
           REGION "SEND TO HMI"
               #saveAct := #partCall.row[#i].pbSelection.actuate;
               #partCall.row[#i] := #requests.row[#pRow];
               #partCall.row[#i].pbSelection.actuate := #saveAct;
           END_REGION

       END_FOR;
   END_REGION
END_FUNCTION_BLOCK

FUNCTION_BLOCK "Clear Part Requests"   // FB17, SCL
{ S7_Optimized_Access := 'TRUE' }
VERSION : 0.1
   VAR_INPUT
      clearRequest : Bool;
   END_VAR
   VAR_IN_OUT
      requests : "Part Request Data";
      partCall : "Part Call Screen";
      currentRowCount : Int;
   END_VAR
   VAR_TEMP
      blankRow : "Table Row";
      i : Int;
      maxRows : Int;
   END_VAR
BEGIN
   REGION "ON REQUEST"
       IF #clearRequest THEN

           REGION "HMI TABLE"

               REGION "COPY TO LOCAL"
                   #maxRows := "partReqHmiRowCount";
               END_REGION

               REGION "CLEAR ROWS"
                   FOR #i := 0 TO #maxRows DO
                       #partCall.row[#i] := #blankRow;
                   END_FOR;
               END_REGION

           END_REGION

           REGION "PART REQUEST DATA BASE"

               REGION "COPY TO LOCAL"
                   #maxRows := "partReqDataRowCount";
               END_REGION

               REGION "CLEAR ROWS"
                   FOR #i := 0 TO #maxRows DO
                       #requests.row[#i] := #blankRow;
                       #currentRowCount := 0;
                   END_FOR;
               END_REGION

           END_REGION

       END_IF;
   END_REGION
END_FUNCTION_BLOCK

FUNCTION_BLOCK "Load Default Timer Presets"   // FB18, SCL
{ S7_Optimized_Access := 'TRUE' }
VERSION : 0.1
   VAR_INPUT
      req : Bool;
   END_VAR
   VAR_IN_OUT
      stations : "Stations";
   END_VAR
   VAR
      oldReq : Bool;
   END_VAR
   VAR_TEMP
      alotted : Real;
      btnCount : Int;
      critical : Real;
      i : Int;
      j : Int;
      partNumber : WString;
      stnCount : Int;
      tmrReal : Real;
   END_VAR
BEGIN
   REGION "COPY TO LOCAL"
       #alotted := "defaultAlotted";
       #btnCount := "ptsPerStn";
       #critical := "defaultCritical";
       #stnCount := #stnCount;
   END_REGION

   REGION "ON REQUEST RISING EDGE"
       IF #req AND NOT #oldReq THEN

           REGION "LOOP THROUGH STATIONS" 
               FOR #i := 0 TO #stnCount DO

                   REGION "LOOP THROUGH BUTTONS"
                       FOR #j := 0 TO #btnCount DO

                           REGION "COPY TO LOCAL"
                               #partNumber := #stations.me[#i].partNumbers[#j];
                           END_REGION

                           REGION "IF BUTTON HAS ASSOCIATED PN"
                               IF LEN(#partNumber) <> 0 THEN

                                   REGION "COPY TO LOCAL"
                                       #tmrReal := #stations.me[#i].presetTime.allotted[#j];
                                   END_REGION

                                   REGION "ON NO TIME ENTERED"
                                       IF #tmrReal = 0.0 THEN

                                           REGION "ASSIGN ALLOTTED VALUES"
                                               #stations.me[#i].presetTime.allotted[#j] := #alotted;
                                           END_REGION

                                       END_IF;
                                   END_REGION

                                   REGION "COPY TO LOCAL"
                                       #tmrReal := #stations.me[#i].presetTime.critical[#j];
                                   END_REGION

                                   REGION "ON NO TIME ENTERED"
                                       IF #tmrReal = 0.0 THEN

                                           REGION "ASSIGN CRITICAL VALUES"
                                               #stations.me[#i].presetTime.critical[#j] := #critical;
                                           END_REGION

                                       END_IF;
                                   END_REGION

                               END_IF;
                           END_REGION

                       END_FOR;
                   END_REGION

               END_FOR;
           END_REGION

       END_IF;
   END_REGION

   REGION "CHANGE DETECTION"
       #oldReq := #req;
   END_REGION ;
END_FUNCTION_BLOCK

FUNCTION_BLOCK "LED Populate Sign"   // FB19, SCL
{ S7_Optimized_Access := 'TRUE' }
VERSION : 0.1
   VAR_INPUT
      requests : "Part Request Data";
   END_VAR
   VAR_IN_OUT
      ledData : "LED Sign Data";
   END_VAR
   VAR_TEMP
      animate : USInt;
      i : Int;
      visibleRows : Int;
      tempRow : "Table Row";
   END_VAR
BEGIN
   REGION "COPY TO LOCAL"
       #visibleRows := "ledRowCount";
   END_REGION

   REGION "POPULATE SIGN DATA"

       REGION "FOR EACH ROW ON SIGN"
           FOR #i := 0 TO #visibleRows DO

               REGION "GET ROW"
                   #tempRow := #requests.row[#i];
               END_REGION

               REGION "LINE LABEL DARK MODE"                
                   "Dark Mode"(#tempRow.tfLine.animate);
               END_REGION

               REGION "DROP ZONE DARK MODE"
                   "Dark Mode"(#tempRow.tfDropZone.animate);
               END_REGION

               REGION "PART NUMBER DARK MODE"

                   REGION "SINGLE LINE"
                       "Dark Mode"(#tempRow.tfPartNumber.animateSL);
                   END_REGION

                   REGION "DOUBLE LINE"
                       "Dark Mode"(#tempRow.tfPartNumber.animateDL);
                   END_REGION

               END_REGION

               REGION "TIME DARK MODE"
                   "Dark Mode"(#tempRow.tfTime.animate);
               END_REGION

               REGION "SEND TO SIGN"
                   #ledData.row[#i] := #tempRow;
               END_REGION

           END_FOR;
       END_REGION

   END_REGION
END_FUNCTION_BLOCK

FUNCTION_BLOCK "Station Selection"   // FB20, SCL
{ S7_Optimized_Access := 'TRUE' }
VERSION : 0.1
   VAR_IN_OUT
      settings : "Settings";
      stations : "Stations";
   END_VAR
   VAR
      firstStn : Int;
      rt : "Runtime Data";
      selectionExe : Bool;
      old : Struct
         prevGrp : Bool;
         nextGrp : Bool;
         stnSlct : Array[0..11] of Bool;
      END_STRUCT;
   END_VAR
   VAR_TEMP
      animate : USInt;
      btnPress : Bool;
      count : Int;
      currentBtn : Bool;
      evalObjCount : Int;
      i : Int;
      oldBtn : Bool;
      pStn : Int;
      stnCount : Int;
      stnName : WString;
      stnSelected : Bool;
      selState : Bool;
      selStnCount : Int;
      timerExpired : Bool;
      stnSelLblCount : Int;
   END_VAR
   VAR CONSTANT
      ptTimer : Real := 1.5;
   END_VAR
BEGIN
   REGION "UI INTERACTION ANIMATIONS"

       REGION "NEXT GROUP"
           #btnPress := #settings.stations.nextGroup.actuate;
           #animate := "Animate Bool"(colorTrue := "BgLGr",
                                      colorFalse := "BgGray",
                                      evalSignal := #btnPress);
           #settings.stations.nextGroup.animate := #animate;
       END_REGION

       REGION "PREVIOUS GROUP"
           #btnPress := #settings.stations.prevGroup.actuate;
           #animate := "Animate Bool"(colorTrue := "BgLGr",
                                      colorFalse := "BgGray",
                                      evalSignal := #btnPress);
           #settings.stations.prevGroup.animate := #animate;
       END_REGION

       REGION "SELECT ALL STATIONS"
           #btnPress := #settings.stations.selectAll.actuate;
           #animate := "Animate Bool"(colorTrue := "BgLGr",
                                      colorFalse := "BgGray",
                                      evalSignal := #settings.stations.selectAll.actuate);
           #settings.stations.selectAll.animate := #animate;
       END_REGION

   END_REGION

   REGION "POPULATE STATION LABELS"

       REGION "PROCESS NEXT GROUP PRESS"

           REGION "COPY TO LOCAL"
               #stnCount := #stnCount;
               #currentBtn := #settings.stations.nextGroup.actuate;
               #oldBtn := #old.nextGrp;
           END_REGION

           REGION "FALLING EDGE OF NEXT GROUP"
               IF NOT #currentBtn AND #oldBtn THEN

                   REGION "INCREMENT FIRST STATION"
                       #firstStn := #firstStn + 2;
                   END_REGION

                   REGION "UPPER LIMIT ROLL OVER"
                       IF #firstStn > #stnCount THEN
                           #firstStn := #firstStn - #stnCount - 1;
                       END_IF;
                   END_REGION

               END_IF;
           END_REGION

           REGION "NEXT GROUP CHANGE DETECTION"
               #old.nextGrp := #currentBtn;
           END_REGION

       END_REGION

       REGION "PROCESS PREVIOUS GROUP PRESS"

           REGION "COPY TO LOCAL"
               #currentBtn := #settings.stations.prevGroup.actuate;
               #oldBtn := #old.prevGrp;
               #stnCount := #stnCount;
           END_REGION

           REGION "FALLING EDGE OF PREVIOUS GROUP"
               IF NOT #currentBtn AND #oldBtn THEN

                   REGION "DECREMENT FIRST STATION"
                       #firstStn := #firstStn - 2;
                   END_REGION

                   REGION "LOWER LIMIT ROLL OVER"
                       IF #firstStn < 0 THEN
                           #firstStn := #firstStn + #stnCount + 1;
                       END_IF;
                   END_REGION

               END_IF;
           END_REGION

           REGION "PREVIOUS GROUP CHANGE DETECTION"
               #old.prevGrp := #currentBtn;
           END_REGION

       END_REGION

       REGION "WRITE LABEL"

           REGION "COPY TO LOCAL"
               #evalObjCount := "hmiSelStnCount";
               #stnCount := "stnCount";
           END_REGION

           REGION "FOR EACH STATION SELECTION BUTTON"
               FOR #i := 0 TO #evalObjCount DO

                   REGION "CALCULATE POINTER"
                       #pStn := #firstStn + #i;
                   END_REGION

                   REGION "UPPER LIMIT ROLL OVER"
                       IF #pStn > #stnCount THEN
                           #pStn := #firstStn + #i - #stnCount - 1;
                       END_IF;
                   END_REGION

                   REGION "BUILD NAME"
                       #stnName := CONCAT_WSTRING(IN1 := #stations.me[#pStn].line,
                                                  IN2 := wstring#' ',
                                                  IN3 := "Strip Sign"(USINT_TO_WSTRING(#stations.me[#pStn].dropZone)));
                   END_REGION

                   REGION "WRITE NAME"
                       #settings.stations.selectBtns[#i].label := #stnName;
                   END_REGION

               END_FOR;
           END_REGION

       END_REGION

   END_REGION

   REGION "SINGLE STATION SELECTION"

       REGION "COPY TO LOCAL"
           #stnSelLblCount := "hmiSelStnCount";
       END_REGION

       REGION "LOOP THROUGH DISPLAYED STATIONS"
           FOR #i := 0 TO #stnSelLblCount DO

               REGION "CALCULATE POINTER"
                   #pStn := #firstStn + #i;
               END_REGION

               REGION "UPPER LIMIT ROLL OVER"
                   #stnCount := "stnCount";
                   IF #pStn > #stnCount THEN
                       #pStn := #firstStn + #i - #stnCount - 1;
                   END_IF;
               END_REGION

               REGION "COPY TO LOCAL"
                   #currentBtn := #settings.stations.selectBtns[#i].actuate;
                   #oldBtn := #old.stnSlct[#i];
               END_REGION

               REGION "TOGGLE STATE ON FALLING EDGE"
                   IF NOT #currentBtn AND #oldBtn THEN
                       #selState := #stations.me[#pStn].settings.selected;
                       #selState := NOT #selState;
                       #stations.me[#pStn].settings.selected := #selState;
                   END_IF;
               END_REGION

               REGION "STATION SELECTION CHANGE DETECTION"
                   #old.stnSlct[#i] := #currentBtn;
               END_REGION

           END_FOR;
       END_REGION

   END_REGION

   REGION "MULTI SELECT TIMER"

       REGION "RUNTIME CALL"
           #rt.elapsed := RUNTIME(#rt.mem);
       END_REGION

       REGION "TIMER"

           REGION "COPY TO LOCAL"
               #btnPress := #settings.stations.selectAll.actuate;
           END_REGION

           REGION "ACCUMULATE RT VALUES"
               IF #btnPress THEN
                   #rt.asReal += LREAL_TO_REAL(#rt.elapsed);
               END_IF;
           END_REGION

           REGION "SET TIMER FLAG"
               IF #rt.asReal < #ptTimer THEN
                   #timerExpired := FALSE;
               END_IF;
               IF #rt.asReal >= #ptTimer THEN
                   #timerExpired := TRUE;
                   #rt.asReal := 0.0;
               END_IF;
           END_REGION

           REGION "RESET ACCUMULATED VALUE"
               IF NOT #btnPress THEN
                   #rt.asReal := 0.0;
                   #selectionExe := FALSE;
               END_IF;
           END_REGION

       END_REGION

   END_REGION

   REGION "EVALUATE MULTI SELECTION"
       IF #timerExpired AND NOT #selectionExe THEN

           REGION "COPY TO LOCAL"
               #selStnCount := #settings.stations.selCount;
           END_REGION

           REGION "SELECT ALL"
               IF #selStnCount < "stnCount" THEN
                   "Select Stations"(mode := TRUE,
                                     stations := #stations);
               END_IF;
           END_REGION

           REGION "DESELECT ALL"
               IF #selStnCount = "stnCount" THEN
                   "Select Stations"(mode := FALSE,
                                     stations := #stations);
               END_IF;
           END_REGION

           REGION "FLAG SELECTION EXECUTED"
               #selectionExe := TRUE;
           END_REGION

       END_IF;
   END_REGION

   REGION "SELECTION ANIMATIONS"

       REGION "COPY TO LOCAL"
           #stnSelLblCount := "hmiSelStnCount";
           #stnCount := "stnCount";
       END_REGION

       REGION "LOOP THROUGH BUTTONS"
           FOR #i := 0 TO #stnSelLblCount DO

               REGION "CALCULATE POINTER"
                   #pStn := #firstStn + #i;
               END_REGION

               REGION "UPPER LIMIT ROLL OVER"
                   IF #pStn > #stnCount THEN
                       #pStn := #firstStn + #i - #stnCount - 1;
                   END_IF;
               END_REGION

               REGION "COPY TO LOCAL"
                   #currentBtn := #settings.stations.selectBtns[#i].actuate;
                   #stnSelected := #stations.me[#pStn].settings.selected;
               END_REGION

               REGION "DRAW SELCTION HIGHLIGHTS"
                   #animate := "Animate Bool"(colorTrue := "BgLTe",
                                              colorFalse := "BgGray",
                                              evalSignal := #stnSelected);
               END_REGION

               REGION "ANIMATE BUTTON PRESS"
                   #animate := "Animate Bool"(colorTrue := "BgDTe",
                                              colorFalse := #animate,
                                              evalSignal := #currentBtn);
                   #settings.stations.selectBtns[#i].animate := #animate;
               END_REGION

           END_FOR;
       END_REGION

   END_REGION

   REGION "COUNT SELECTED STATIONS"

       REGION "INITIALIZE LOCAL"
           #count := 0;
           #evalObjCount := "stnCount";
       END_REGION

       REGION "LOOP THROUGH STATIONS"
           FOR #i := 0 TO #evalObjCount DO

               REGION "INCREMENT COUNT ON SELECTION"
                   #stnSelected := #stations.me[#i].settings.selected;
                   IF #stnSelected THEN
                       #count += 1;
                   END_IF;
               END_REGION

           END_FOR;
       END_REGION

       REGION "SAVE COUNT"
           #settings.stations.selCount := #count;
       END_REGION

   END_REGION
END_FUNCTION_BLOCK

FUNCTION_BLOCK "KP8 Button Selections"   // FB21, SCL
{ S7_Optimized_Access := 'TRUE' }
VERSION : 0.1
   VAR_INPUT
      reset : Bool;
   END_VAR
   VAR_IN_OUT
      settings : "Settings";
      stations : "Stations";
   END_VAR
   VAR
      enableState : Bool;
      oldBtnPresses : Array[0..7] of Bool;
      oldSelState : Array[0..7] of Bool;
      oldSelStnCount : Int;
      rt : "Runtime Data";
      timerExpired : Bool;
      selectionExe : Bool;
   END_VAR
   VAR_TEMP
      animate : USInt;
      btnCount : Int;
      btnPress : Bool;
      count : Int;
      i : Int;
      j : Int;
      mode : Bool;
      oldPress : Bool;
      pBtn : Int;
      selBtnCount : Int;
      selStnCount : Int;
      stnCount : Int;
      stnSelected : Bool;
   END_VAR
   VAR CONSTANT
      selectAllTime : Real := 1.5;
   END_VAR
BEGIN
   REGION "ENABLE KP8 BUTTON ASSIGNMENT SECTION"

       REGION "ENABLE"

           REGION "COPY TO LOCAL"
               #selStnCount := #settings.stations.selCount;
           END_REGION

           REGION "ON CHANGE IN SELECTED STATION COUNT"
               IF #selStnCount <> 0 AND #selStnCount <> #oldSelStnCount THEN

                   REGION "ENABLE KP8 SELECTIONS"
                       #enableState := TRUE;
                   END_REGION

               END_IF;
           END_REGION

       END_REGION

       REGION "DISABLE"

           REGION "COPY TO LOCAL"
               #selStnCount := #settings.stations.selCount;
               #btnCount := "ptsPerStn";
           END_REGION

           REGION "ON DESELETION OF LAST STATION"
               IF #selStnCount = 0 AND #selStnCount <> #oldSelStnCount THEN

                   REGION "RESET ENABLED STATE"
                       #enableState := FALSE;
                   END_REGION

                   REGION "RESET BUTTON SELECTION STATES"
                       FOR #i := 0 TO #btnCount DO
                           #settings.kp8.btnSelState[#i] := FALSE;
                       END_FOR;
                   END_REGION

               END_IF;
           END_REGION

       END_REGION

   END_REGION

   REGION "SINGLE BUTTON SELECTION"

       REGION "COPY TO LOCAL"
           #btnCount := "ptsPerStn";
       END_REGION

       REGION "LOOP THROUGH BUTTONS"
           FOR #i := 0 TO #btnCount DO

               REGION "EXCLUDE STOP RUNTIME AND RESET SELECTED BUTTONS"
                   IF #i <> 0 AND #i <> 4 THEN

                       REGION "COPY TO LOCAL"

                           REGION "CALCULATE BUTTON POINTER"
                               CASE #i OF
                                   1:
                                       #pBtn := 5;
                                   2:
                                       #pBtn := 3;
                                   3:
                                       #pBtn := 1;
                                   5:
                                       #pBtn := 4;
                                   6:
                                       #pBtn := 2;
                                   7:
                                       #pBtn := 0;
                                   ELSE
                                       ;
                               END_CASE;
                           END_REGION

                           #btnPress := #settings.kp8.buttons[#i].actuate OR #settings.viewingStation.btns[#pBtn].select.actuate;
                           #oldPress := #oldBtnPresses[#i];

                       END_REGION

                       REGION "TOGGLE STATE ON FALLING EDGE"
                           IF NOT #btnPress AND #oldPress THEN
                               #settings.kp8.btnSelState[#i] := NOT #settings.kp8.btnSelState[#i];
                               #settings.kp8.selBtnNumber := #i;
                           END_IF;
                       END_REGION

                       REGION "SAVE SELECTED BUTTON NUMBER ON DESELECT"
                           IF NOT #settings.kp8.btnSelState[#i] AND #oldSelState[#i] THEN
                               FOR #j := 0 TO #btnCount DO
                                   IF #settings.kp8.btnSelState[#j] THEN
                                       #settings.kp8.selBtnNumber := #j;
                                   END_IF;
                               END_FOR;
                           END_IF;
                       END_REGION

                       REGION "KP8 BUTON SELECTION CHANGE DETECTION"
                           #oldBtnPresses[#i] := #btnPress;
                       END_REGION

                   END_IF;
               END_REGION

           END_FOR;
       END_REGION

   END_REGION

   REGION "MULTI BUTTON SELECTION"

       REGION "MULTI SELECT TIMER"

           REGION "RUNTIME CALL"
               #rt.elapsed := RUNTIME(#rt.mem);
           END_REGION

           REGION "TIMER"

               REGION "COPY TO LOCAL"
                   #btnPress := #settings.kp8.selectButtons.actuate;
               END_REGION

               REGION "ACCUMULATE RT VALUES"
                   IF #btnPress THEN
                       #rt.asReal += LREAL_TO_REAL(#rt.elapsed);
                   END_IF;
               END_REGION

               REGION "SET TIMER FLAG"
                   IF #rt.asReal < #selectAllTime THEN
                       #timerExpired := FALSE;
                   END_IF;
                   IF #rt.asReal >= #selectAllTime THEN
                       #timerExpired := TRUE;
                       #rt.asReal := 0.0;
                   END_IF;
               END_REGION

               REGION "RESET ACCUMULATED VALUE"
                   IF NOT #btnPress THEN
                       #rt.asReal := 0.0;
                       #selectionExe := FALSE;
                   END_IF;
               END_REGION

           END_REGION

       END_REGION

       REGION "EVALUATE MULTI SELECTION"
           IF #timerExpired AND NOT #selectionExe THEN

               REGION "COPY TO LOCAL"
                   #btnCount := "ptsPerStn";
                   #selBtnCount := #settings.kp8.selCount;
               END_REGION

               REGION "SELECT ALL"
                   IF #selBtnCount < #btnCount - 1 THEN
                       #mode := TRUE;
                   END_IF;
               END_REGION

               REGION "DESELECT ALL"
                   IF #selBtnCount = #btnCount - 1 THEN
                       #mode := FALSE;
                   END_IF;
               END_REGION

               REGION "SAVE SELECTIONS"
                   FOR #i := 0 TO #btnCount DO

                       REGION "EXCLUDE STOP RUNTIME AND RESET SELECTED BUTTONS"
                           IF #i <> 0 AND #i <> 4 THEN

                               REGION "PERFROM SELECTION"
                                   #settings.kp8.btnSelState[#i] := #mode;
                               END_REGION

                           END_IF;
                       END_REGION

                   END_FOR;
               END_REGION

               REGION "SET SELECED BUTTON NUMBER TO 1"
                   #settings.kp8.selBtnNumber := 0;
               END_REGION

               REGION "FLAG SELECTION EXECUTED"
                   #selectionExe := TRUE;
               END_REGION

           END_IF;
       END_REGION
   END_REGION

   REGION "SAVE BUTTON SELECTIONS TO STATIONS"

       REGION "COPY TO LOCAL"
           #selStnCount := #settings.stations.selCount;
       END_REGION

       REGION "ON CHANGE IN BUTTON OR STATION SELECTON"
           IF #settings.kp8.btnSelState <> #oldSelState OR #selStnCount <> #oldSelStnCount THEN

               REGION "COPY TO LOCAL"
                   #stnCount := #stnCount;
               END_REGION

               REGION "FOR SELECTED STATIONS"
                   FOR #i := 0 TO #stnCount DO
                       #stnSelected := #stations.me[#i].settings.selected;
                       IF #stnSelected THEN

                           REGION "SAVE BUTTON SELECTION STATE"
                               #stations.me[#i].settings.btnSelection := #settings.kp8.btnSelState;
                           END_REGION

                       END_IF;
                   END_FOR;
               END_REGION

           END_IF;
       END_REGION

       REGION "SELECTED STATION COUNT CHANGE DETECTION"
           #oldSelStnCount := #selStnCount; 
       END_REGION

   END_REGION

   REGION "COUNT SELECTED BUTTONS"

       REGION "COPY TO LOCAL"
           #btnCount := "ptsPerStn";
       END_REGION 

       REGION "ON CHANGE IN BUTTON SELECTION STATES"
           IF #settings.kp8.btnSelState <> #oldSelState THEN

               REGION "INITIALIZE LOCAL"
                   #count := 0;
               END_REGION

               REGION "FOR EACH SELECTED BUTTON"
                   FOR #i := 0 TO #btnCount DO
                       IF #settings.kp8.btnSelState[#i] THEN

                           REGION "INCREMENT COUNT"
                               #count := #count + 1;
                           END_REGION

                       END_IF;
                   END_FOR;
               END_REGION

               REGION "SAVE COUNT"
                   #settings.kp8.selCount := #count;
               END_REGION

           END_IF;
       END_REGION

   END_REGION 

   REGION "UI INTERACTION ANIMATIONS"

       REGION "SELECT ALL BUTTONS"
           #btnPress := #settings.kp8.selectButtons.actuate;
           #animate := "Animate Bool"(colorTrue := "BgLGr",
                                      colorFalse := "BgGray",
                                      evalSignal := #btnPress);
           #settings.kp8.selectButtons.animate := #animate;
       END_REGION

       REGION "STOP RESET SELECTED STATION"
           #btnPress := #settings.kp8.buttons[0].actuate;
           #animate := "Animate Bool"(colorTrue := "FgGray",
                                      colorFalse := "BgGray",
                                      evalSignal := #btnPress);
           #settings.kp8.buttons[0].animate := #animate;
       END_REGION

       REGION "STOP RUNTIME"
           #btnPress := #settings.kp8.buttons[4].actuate;
           #animate := "Animate Bool"(colorTrue := "FgGray",
                                      colorFalse := "BgGray",
                                      evalSignal := #btnPress);
           #settings.kp8.buttons[4].animate := #animate;
       END_REGION

       REGION "BUTTON SELECTIONS"

           REGION "COPY TO LOCAL"
               #btnCount := "ptsPerStn";
           END_REGION

           REGION "FOR EACH BUTTON"     
               FOR #i := 0 TO #btnCount DO

                   REGION "EXCLUDE STOP RUNTIME AND RESET SELECTED BUTTONS"
                       IF #i <> 0 AND #i <> 4 THEN

                           REGION "ANIMATE"

                               REGION "COPY TO LOCAL"
                                   #btnPress := #settings.kp8.buttons[#i].actuate;
                               END_REGION

                               REGION "ENABLE/DISABLE"
                                   #animate := "Animate Bool"(colorTrue := "BgGray",
                                                              colorFalse := "disabled",
                                                              evalSignal := #enableState);
                               END_REGION

                               REGION "ENABLED SUB ANIMATIONS"
                                   IF #enableState THEN

                                       REGION "BUTTON SELECTED"
                                           #animate := "Animate Bool"(colorTrue := "BgLTe",
                                                                      colorFalse := #animate,
                                                                      evalSignal := #settings.kp8.btnSelState[#i]);
                                       END_REGION

                                       REGION "BUTTON UP/DOWN"
                                           #animate := "Animate Bool"(colorTrue := "BgDTe",
                                                                      colorFalse := #animate,
                                                                      evalSignal := #btnPress);
                                       END_REGION
                                   END_IF;
                               END_REGION

                               REGION "SAVE ANIMATION"
                                   #settings.kp8.buttons[#i].animate := #animate;
                               END_REGION

                           END_REGION

                       END_IF;
                   END_REGION

               END_FOR;
           END_REGION

       END_REGION

   END_REGION

   REGION "DRAW KP8 BUTTON LABELS"
       IF #reset THEN
           #settings.kp8.buttons[1].label := wstring#'6';
           #settings.kp8.buttons[2].label := wstring#'4';
           #settings.kp8.buttons[3].label := wstring#'2';
           #settings.kp8.buttons[5].label := wstring#'5';
           #settings.kp8.buttons[6].label := wstring#'3';
           #settings.kp8.buttons[7].label := wstring#'1';
       END_IF;
   END_REGION

   REGION "CHANGE DETECTION"
       #oldSelState := #settings.kp8.btnSelState;
   END_REGION
END_FUNCTION_BLOCK

FUNCTION_BLOCK "Buffer Log: Part Requests"   // FB22, SCL
{ S7_Optimized_Access := 'TRUE' }
VERSION : 0.1
   VAR_INPUT
      stations : "Stations";
   END_VAR
   VAR_IN_OUT
      logBuffer : "Part Req Log";
      logFlag : Int;
   END_VAR
   VAR
      clpsLogTime : Real;
      old : Struct
         ordered : "Station Old Presses";
         requested : "Station Old Presses";
      END_STRUCT;
      pLogBuffer : Int;
      rt : "Runtime Data";
   END_VAR
   VAR_TEMP
      address : Int;
      btnCount : Int;
      clpsFlag : Bool;
      i : Int;
      j : Int;
      oldPartOrdered : Bool;
      oldPartReq : Bool;
      partOrdered : Bool;
      partReq : Bool;
      stnCount : Int;
      readTimeRetVal : Int;
      blankRow : "Part Req Log Row";
   END_VAR
   VAR CONSTANT
      clpsItrvl : Real := 2.0;
      fulfilled : Int := 3;
      ordered : Int := 2;
      requested : Int := 1;
   END_VAR
BEGIN
   REGION "RUNTIME CALL"
       #rt.elapsed := RUNTIME(#rt.mem);
       #rt.asReal := LREAL_TO_REAL(#rt.elapsed);
   END_REGION

   REGION "COPY TO LOCAL"
       #btnCount := "ptsPerStn";
       #stnCount := "stnCount";
   END_REGION

   REGION "FOR EACH STATION"
       FOR #i := 0 TO #stnCount DO

           REGION "FOR EACH BUTTON"
               FOR #j := 0 TO #btnCount DO

                   REGION "COPY TO LOCAL"
                       #partOrdered := #stations.me[#i].partOrdered[#j];
                       #partReq := #stations.me[#i].partRequested[#j];
                       #oldPartOrdered := #old.ordered.me[#i,#j];
                       #oldPartReq := #old.requested.me[#i,#j];
                   END_REGION;

                   REGION "CALCULATE ADDRESS"
                       #address := (#i + 1) * 10 + #j + 1;
                   END_REGION

                   REGION "ON PART REQUEST RISING EDGE"
                       IF #partReq AND NOT #oldPartReq THEN

                           REGION "LOG ENTRY"
                               #logBuffer.me[#pLogBuffer] := "Buffer Part Req Log Row: Generate"(address := #address,
                                                                                        type := #requested);
                           END_REGION

                           REGION "INCREMENT POINTER"
                               #pLogBuffer += 1;
                           END_REGION

                       END_IF;
                   END_REGION

                   REGION "ON PART ORDERED RISING EDGE"
                       IF #partOrdered AND NOT #oldPartOrdered THEN

                           REGION "REQUEST TYPE"
                               #logBuffer.me[#pLogBuffer] := "Buffer Part Req Log Row: Generate"(address := #address,
                                                                                                 type := #ordered);
                           END_REGION

                           REGION "INCREMENT POINTER"
                               #pLogBuffer += 1;
                           END_REGION

                       END_IF;
                   END_REGION

                   REGION "ON PART REQUEST FALLING EDGE"
                       IF NOT #partReq AND #oldPartReq THEN

                           REGION "REQUEST TYPE"
                               #logBuffer.me[#pLogBuffer] := "Buffer Part Req Log Row: Generate"(
                                   address := #address,
                                   type := #fulfilled
                               );
                           END_REGION

                           REGION "INCREMENT POINTER"
                               #pLogBuffer += 1;
                           END_REGION

                       END_IF;
                   END_REGION

                   REGION "SAVE FOR CHANGE DETECTION"
                       #old.requested.me[#i, #j] := #partReq;
                       #old.ordered.me[#i, #j] := #partOrdered;
                   END_REGION

               END_FOR;
           END_REGION

       END_FOR;
   END_REGION

   REGION "SEND TO HMI"

       REGION "ON ENTRY IN BUFFER"
           IF #logBuffer.me[0].address <> 0 THEN

               REGION "TIMER"
                   #clpsLogTime += #rt.asReal;
                   IF #clpsLogTime >= #clpsItrvl THEN
                       #clpsLogTime := 0.0;
                       #clpsFlag := TRUE;
                   END_IF;
               END_REGION

               REGION "EXECUTE COLLAPSE"
                   IF #clpsFlag THEN

                       REGION "MOVE BUFFER UP ONE POSITION"
                           FOR #i := 0 TO 98 DO
                               #logBuffer.me[#i] := #logBuffer.me[#i + 1];
                           END_FOR;
                       END_REGION

                       REGION "DELETE LAST ROW"
                           #logBuffer.me[99] := #blankRow;
                       END_REGION

                       REGION "FLAG FOR HMI"
                           #logFlag += 1;
                           IF #logFlag > 9 THEN
                               #logFlag := 0;
                           END_IF;
                       END_REGION

                       REGION "DECREMENT POINTER"
                           #pLogBuffer -= 1;
                       END_REGION

                   END_IF;
               END_REGION

           END_IF;
       END_REGION

   END_REGION

   REGION "RESET TIMER"
       IF #logBuffer.me[0].address = 0 THEN
           #clpsLogTime := 0.0;
       END_IF;
   END_REGION
END_FUNCTION_BLOCK

FUNCTION_BLOCK "Enable Assignment Pair"   // FB23, SCL
{ S7_Optimized_Access := 'TRUE' }
VERSION : 0.1
   VAR_INPUT
      disable : Bool;
      enable : Bool;
   END_VAR
   VAR_IN_OUT
      value : WString;
      assignAnimate : USInt;
      ioFieldAnimate : USInt;
   END_VAR
   VAR
      old : Struct
         disabled : Bool;
         enabled : Bool;
      END_STRUCT;
   END_VAR
BEGIN
   REGION "DISABLED"    
       IF #disable THEN
           #value := wstring#'';
           #assignAnimate := "disabled";
           #ioFieldAnimate := "disabled";
       END_IF;
   END_REGION

   REGION "ENABLED"
           IF #enable THEN
               #assignAnimate := "BgGray";
               #ioFieldAnimate := "BgWh";
           END_IF;
   END_REGION
END_FUNCTION_BLOCK

FUNCTION_BLOCK "Assign Button Parameters"   // FB24, SCL
{ S7_Optimized_Access := 'TRUE' }
VERSION : 0.1
   VAR_INPUT
      settings : "Settings";
   END_VAR
   VAR_IN_OUT
      stations : "Stations";
   END_VAR
   VAR
      old : Struct
         allotted : Bool;
         critical : Bool;
         pn : Bool;
      END_STRUCT;
   END_VAR
   VAR_TEMP
      assign : Bool;
      btn : Struct
         allotted : Bool;
         critical : Bool;
         pn : Bool;
      END_STRUCT;
      btnCount : Int;
      btnSelected : Bool;
      i : Int;
      j : Int;
      partNumber : WString;
      stnCount : Int;
      stnSelected : Bool;
      timerReal : Real;
   END_VAR
BEGIN
   REGION "COPY TO LOCACL"
       #stnCount := "stnCount";
       #btnCount := "ptsPerStn";
       #btn.allotted := #settings.alotted.assign.actuate;
       #btn.critical := #settings.critical.assign.actuate;
       #btn.pn := #settings.partNumber.assign.actuate;
   END_REGION

   REGION "ASSIGNMENT PULSE"
       #assign := (#btn.allotted AND NOT #old.allotted)
                   OR (#btn.critical AND NOT #old.critical)
                   OR (#btn.pn AND NOT #old.pn);
   END_REGION

   REGION "ON ASSIGNMENT PULSE"
       IF #assign THEN

           REGION "PROCESS VARIABLE"

               REGION "PART NUMBER"
                   IF #btn.pn THEN
                       #partNumber := #settings.partNumber.ioField.value;
                   END_IF;
               END_REGION

               REGION "CRITICAL TIME"
                   IF #btn.critical THEN
                       #timerReal := "WString Timer to Real"(#settings.critical.ioField.value);
                   END_IF;
               END_REGION

               REGION "ALLOTTED TIME"
                   IF #btn.allotted THEN
                       #timerReal := "WString Timer to Real"(#settings.alotted.ioField.value);
                   END_IF;
               END_REGION

           END_REGION

           REGION "FOR EACH STATION"
               FOR #i := 0 TO #stnCount DO

                   REGION "COPY TO LOCAL"
                       #stnSelected := #stations.me[#i].settings.selected;
                   END_REGION

                   REGION "ON SELECTED STATION"
                       IF #stnSelected THEN

                           REGION "FOR EACH BUTTON"
                               FOR #j := 0 TO #btnCount DO

                                   REGION "COPY TO LOCAL"
                                       #btnSelected := #stations.me[#i].settings.btnSelection[#j];
                                   END_REGION

                                   REGION "ON SELECTED BUTTON"
                                       IF #btnSelected THEN

                                           REGION "ASSIGN PART NUMBER"
                                               IF #btn.pn THEN
                                                   #stations.me[#i].partNumbers[#j] := #partNumber;
                                               END_IF;
                                           END_REGION

                                           REGION "ASSIGN ALLOTTED TIME"
                                               IF #btn.allotted THEN
                                                   #stations.me[#i].presetTime.allotted[#j] := #timerReal;
                                               END_IF;
                                           END_REGION

                                           REGION "ASSIGN CRITICAL TIME"
                                               IF #btn.critical THEN
                                                   #stations.me[#i].presetTime.critical[#j] := #timerReal;
                                               END_IF;
                                           END_REGION

                                       END_IF;
                                   END_REGION

                               END_FOR;
                           END_REGION

                       END_IF;
                   END_REGION

               END_FOR;
           END_REGION

       END_IF;
   END_REGION

   REGION "CHANGE DETECTION"
       #old := #btn;
   END_REGION
END_FUNCTION_BLOCK

FUNCTION_BLOCK "Animate: PN & Timers"   // FB25, SCL
{ S7_Optimized_Access := 'TRUE' }
VERSION : 0.1
   VAR_INPUT
      stations : "Stations";
   END_VAR
   VAR_IN_OUT
      settings : "Settings";
   END_VAR
   VAR
      instPNEntEnable : "Enable Assignment Pair";
      instAlltEntEnable : "Enable Assignment Pair";
      instCrtEntEnable : "Enable Assignment Pair";
   END_VAR
   VAR_TEMP
      animate : USInt;
      disable : Bool;
      enable : Bool;
      selBtnCount : Int;
      selStnCount : Int;
   END_VAR
BEGIN
   REGION "COPY TO LOCAL"
       #selBtnCount := #settings.kp8.selCount;
       #selStnCount := #settings.stations.selCount;
   END_REGION

   REGION "ENABLE/DISABLE FOR PN AND TIMERS"

       REGION "SET DISABLE"
           IF #selStnCount = 0 OR #selBtnCount = 0 THEN
               #disable := TRUE;
               #enable := FALSE;
           END_IF;
       END_REGION

       REGION "SET ENABLE"
           IF #selStnCount <> 0 AND #selBtnCount <> 0 THEN
               #disable := FALSE;
               #enable := TRUE;
           END_IF;
       END_REGION

   END_REGION

   REGION "PN ANIMATION FUNCTIONS"
       #animate := #settings.partNumber.assign.animate;
       #instPNEntEnable(disable := #disable,
                        enable := #enable,
                        value := #settings.partNumber.ioField.value,
                        assignAnimate := #animate,
                        ioFieldAnimate := #settings.partNumber.ioField.animate);
       #animate := "Animate Bool"(colorTrue := "BgLGr",
                                  colorFalse := #animate,
                                  evalSignal := #settings.partNumber.assign.actuate);
       #settings.partNumber.assign.animate := #animate;
   END_REGION

   REGION "ALLOTTED TIME ANIMATION FUNCTIONS"
       #animate := #settings.alotted.assign.animate;
       #instAlltEntEnable(disable := #disable,
                          enable := #enable,
                          value := #settings.alotted.ioField.value,
                          assignAnimate := #animate,
                          ioFieldAnimate := #settings.alotted.ioField.animate);
       #animate := "Animate Bool"(colorTrue := "BgLGr",
                                  colorFalse := #animate,
                                  evalSignal := #settings.alotted.assign.actuate);
       #settings.alotted.assign.animate := #animate;
   END_REGION

   REGION "CRITICAL TIME ANIMATION FUNCTIONS"
       #animate := #settings.critical.assign.animate;
       #instCrtEntEnable(disable := #disable,
                         enable := #enable,
                         value := #settings.critical.ioField.value,
                         assignAnimate := #animate,
                         ioFieldAnimate := #settings.critical.ioField.animate);
       #animate := "Animate Bool"(colorTrue := "BgLGr",
                                  colorFalse := #animate,
                                  evalSignal := #settings.critical.assign.actuate);
       #settings.critical.assign.animate := #animate;
   END_REGION
END_FUNCTION_BLOCK

FUNCTION_BLOCK "Global to Sim"   // FB26, SCL
{ S7_Optimized_Access := 'TRUE' }
VERSION : 0.1
   VAR_INPUT
      stations : "Stations";
   END_VAR
   VAR_IN_OUT
      simStations : "Simulated Stations";
   END_VAR
   VAR
      old : Struct
         nextGrp : Bool;
         prevGrp : Bool;
      END_STRUCT;
   END_VAR
   VAR_TEMP
      animate : USInt;
      btnCount : Int;
      currentBtn : Bool;
      dzLabel : WString;
      firstStn : Int;
      i : Int;
      intBox : Int;
      j : Int;
      kp8Color : DWord;
      label : WString;
      oldBtn : Bool;
      pSim : Int;
      pStn : Int;
      simKP8Count : Int;
      stnCount : Int;
   END_VAR
   VAR CONSTANT
      space : WString := WSTRING#' ';
      lead0 : WString := WSTRING#'0';
      volvo16 : WString := WSTRING#'VOLVO 16';
   END_VAR
BEGIN
   REGION "COPY TO LOCAL"
       #btnCount := "ptsPerStn";
       #firstStn := #simStations.firstStn;
       #stnCount := "stnCount";
       #simKP8Count := "simKP8Count";
   END_REGION

   REGION "RESOLVE STATION POINTER"

       REGION "PROCESS NEXT GROUP PRESS"

           REGION "COPY TO LOCAL"
               #currentBtn := #simStations.down.actuate;
               #oldBtn := #old.nextGrp;
           END_REGION

           REGION "FALLING EDGE OF NEXT GROUP"
               IF NOT #currentBtn AND #oldBtn THEN

                   REGION "INCREMENT FIRST STATION"
                       #firstStn += #simKP8Count;
                   END_REGION

                   REGION "UPPER LIMIT ROLL OVER"
                       IF #firstStn > #stnCount THEN
                           #firstStn -= #stnCount + 1;
                       END_IF;
                   END_REGION

               END_IF;
           END_REGION

           REGION "NEXT GROUP CHANGE DETECTION"
               #old.nextGrp := #currentBtn;
           END_REGION

       END_REGION

       REGION "PROCESS PREVIOUS GROUP PRESS"

           REGION "COPY TO LOCAL"
               #currentBtn := #simStations.up.actuate;
               #oldBtn := #old.prevGrp;
           END_REGION

           REGION "FALLING EDGE OF PREVIOUS GROUP"
               IF NOT #currentBtn AND #oldBtn THEN

                   REGION "DECREMENT FIRST STATION"
                       #firstStn -= #simKP8Count;
                   END_REGION

                   REGION "LOWER LIMIT ROLL OVER"
                       IF #firstStn < 0 THEN
                           #firstStn += #stnCount + 1;
                       END_IF;
                   END_REGION

               END_IF;
           END_REGION

           REGION "PREVIOUS GROUP CHANGE DETECTION"
               #old.prevGrp := #currentBtn;
           END_REGION

       END_REGION

   END_REGION

   REGION "FOR EACH BUTTON"
       FOR #i := 0 TO 11 DO

           REGION "CALCULATE POINTER"
               #pStn := #i + #firstStn;
               #pSim := #i;
           END_REGION

           REGION "UPPER LIMIT ROLL OVER"
               IF #pStn > #stnCount THEN
                   #pStn := #firstStn + #i - #stnCount - 1;
               END_IF;
           END_REGION

           REGION "COPY TO LOCAL"
               #kp8Color := #stations.me[#pStn].kp8Out;
           END_REGION

           REGION "LABEL STATIONS"

               REGION "DETERMINE LINE LABEL"
                   #label := #stations.me[#pStn].line;
                   IF #label = #volvo16 THEN
                       #label := WSTRING#'V16';
                   END_IF;
               END_REGION

               REGION "DETERMINE DROP ZONE LABEL"
                   #intBox := USINT_TO_INT(#stations.me[#pStn].dropZone);
                   IF #intBox <= 9 THEN
                       #dzLabel := CONCAT_WSTRING(IN1 := #lead0,
                                                  IN2 := "Strip Sign"(INT_TO_WSTRING(#intBox)));
                   END_IF;
                   IF #intBox >= 10 THEN
                       #dzLabel := "Strip Sign"(INT_TO_WSTRING(#intBox));
                   END_IF;
               END_REGION

               REGION "WRITE LABEL"
                   #label := CONCAT_WSTRING(IN1 := #label,
                                            IN2 := #space,
                                            IN3 := #dzLabel);
                   #simStations.me[#pSim].stn.label := #label;
               END_REGION

           END_REGION

           REGION "ANIMATE STATION LABEL"
               #simStations.me[#pSim].stn.animate := "BgGray";
           END_REGION

           REGION "FOR EACH BUTTON"
               FOR #j := 0 TO #btnCount DO

                   REGION "COLOR BUTTONS"
                       #animate := "KP8 Color to Sim Animation"(kp8Color := #kp8Color,
                                                                btnNumber := #j);
                       #simStations.me[#pSim].btn.animate[#j] := #animate;
                   END_REGION

                   REGION "WRITE BUTTON LABELS"
                       #intBox := "Pointer Calc: KP8 Labels"(#j);
                       #label := "Strip Sign"(INT_TO_WSTRING(#intBox));
                       #simStations.me[#pSim].btn.labels[#j] := #label;
                   END_REGION

               END_FOR;
           END_REGION

       END_FOR;
   END_REGION

   REGION "SAVE FIRST STATION"
       #simStations.firstStn := #firstStn;
   END_REGION

   REGION "ANIMATE NEXT GROUP PRESS"
       #simStations.down.animate := "Animate Bool"(colorTrue := "BgLGr",
                                                   colorFalse := "BgGray",
                                                   evalSignal := #simStations.down.actuate);
   END_REGION

   REGION "ANIMATE PREV GROUP PARESS"
       #simStations.up.animate := "Animate Bool"(colorTrue := "BgLGr",
                                                 colorFalse := "BgGray",
                                                 evalSignal := #simStations.up.actuate);
   END_REGION
END_FUNCTION_BLOCK

FUNCTION_BLOCK "HMI: Network Health"   // FB31, SCL
{ S7_Optimized_Access := 'TRUE' }
VERSION : 0.1
   VAR_IN_OUT
      ioSystemData : Array[1.."USERDIAG_IO_SYSTEMS_UPPER_LIM"] of "UserDiag_typeIOSystem";
      netHealthScreen : "Network Health Screen";
   END_VAR
   VAR_TEMP
      i : Int;
      animate : Struct
         ok : USInt;
         faulty : USInt;
         lostConn : USInt;
         disabled : USInt;
         problem : USInt;
         wasFaulty : USInt;
         wasLost : USInt;
         wasDisabled : USInt;
         problemGone : USInt;
      END_STRUCT;
   END_VAR
   VAR CONSTANT
      statOk : USInt := 1;
   END_VAR
BEGIN
   #animate.ok := "BgDGr";

   FOR #i := 1 TO "pnioDeviceCount" DO
       #netHealthScreen.pnioDevices[#i].label := #ioSystemData[1].devices[#i].name;
       CASE #ioSystemData[1].devices[#i].state OF
           #statOk:
               #netHealthScreen.pnioDevices[#i].animate := #animate.ok;
           ELSE 
               ;
       END_CASE;
   END_FOR;
END_FUNCTION_BLOCK

FUNCTION_BLOCK "Table Navigatio"   // FB34, SCL
{ S7_Optimized_Access := 'TRUE' }
VERSION : 0.1
   VAR_INPUT
      maxRows : DInt;
      visRows : DInt;
      offset : DInt;
      trigger : Bool;
   END_VAR
   VAR_IN_OUT
      r1 : DInt;
      rowIndices : Array[0..#maxOutRows] of DInt;
   END_VAR
   VAR
      old : Struct
         trigger : Bool := false;
      END_STRUCT;
   END_VAR
   VAR_TEMP
      i : DInt;
      output : Array[0..#maxOutRows] of DInt;
      thisIndex : DInt;
      newR1 : DInt;
   END_VAR
   VAR CONSTANT
      maxOutRows : DInt := 99;
   END_VAR
BEGIN
   IF #trigger AND NOT #old.trigger THEN

       FOR #i := 0 TO #maxOutRows DO
           #output[#i] := -1;
       END_FOR;

       IF #offset > -1000 THEN

           #newR1 := #r1 + #offset;

           IF #newR1 < 0 THEN
               #newR1 := #newR1 + #maxRows;
           END_IF;

           IF #newR1 > #maxRows THEN
               #newR1 := #newR1 - #maxRows;
           END_IF;

       END_IF;

       IF #offset = -1000 THEN
           #newR1 := 0;
       END_IF;

       IF #offset = - 2000 THEN
           #newR1 := #maxRows - #visRows;
       END_IF;

       FOR #i := 0 TO #visRows - 1 DO
           #thisIndex := #newR1 + #i;
           IF #thisIndex < 0 THEN
               #thisIndex := #thisIndex + #maxRows;
           END_IF;
           IF #thisIndex >= #maxRows THEN
               #thisIndex := #thisIndex - #maxRows;
           END_IF;
           #output[#i] := #thisIndex;
       END_FOR;

       #rowIndices := #output;
       #r1 := #newR1;

   END_IF;

   #old.trigger := #trigger;
END_FUNCTION_BLOCK

FUNCTION_BLOCK "KP8 Driver"   // FB101, SCL
{ S7_Optimized_Access := 'FALSE' }
VERSION : 0.1
   VAR_INPUT
      btnIn : Byte;   // byte that contains input data from kp8 buttons
      hardInit : Bool;   // initializes function. can be used for reset
      softInit : Bool;
      btn0Activate : Bool;   // true for on, false for off
      btn0Mode : Bool;   // true for maintained, false for momentary
      btn0Group : Int;
      btn0Flash : Bool;
      btn0ColorOn1 : String[10];   // enter: red OR green OR blue OR yellow OR white OR off
      btn0ColorOn2 : String[10];
      btn0ColorOff : String[10];   // enter: red OR green OR blue OR yellow OR white OR off
      btn1Activate : Bool;   // true for on, false for off
      btn1Mode : Bool;   // true for maintained, false for momentary
      btn1Group : Int;
      btn1Flash : Bool;
      btn1ColorOn1 : String[10];   // enter: red OR green OR blue OR yellow OR white OR off
      btn1ColorOn2 : String[10];
      btn1ColorOff : String[10];   // enter: red OR green OR blue OR yellow OR white OR off
      btn2Activate : Bool;   // true for on, false for off
      btn2Mode : Bool;   // true for maintained, false for momentary
      btn2Group : Int;
      btn2Flash : Bool;
      btn2ColorOn1 : String[10] := '';   // enter: red OR green OR blue OR yellow OR white OR off
      btn2ColorOn2 : String[10];
      btn2ColorOff : String[10];   // enter: red OR green OR blue OR yellow OR white OR off
      btn3Activate : Bool;   // true for on, false for off
      btn3Mode : Bool;   // true for maintained, false for momentary
      btn3Group : Int;
      btn3Flash : Bool;
      btn3ColorOn1 : String[10];   // enter: red OR green OR blue OR yellow OR white OR off
      btn3ColorOn2 : String[10];
      btn3ColorOff : String[10];   // enter: red OR green OR blue OR yellow OR white OR off
      btn4Activate : Bool;   // true for on, false for off
      btn4Mode : Bool;   // true for maintained, false for momentary
      btn4Group : Int;
      btn4Flash : Bool;
      btn4ColorOn1 : String[10];   // enter: red OR green OR blue OR yellow OR white OR off
      btn4ColorOn2 : String[10];
      btn4ColorOff : String[10];   // enter: red OR green OR blue OR yellow OR white OR off
      btn5Activate : Bool;   // true for on, false for off
      btn5Mode : Bool;   // true for maintained, false for momentary
      btn5Group : Int;
      btn5Flash : Bool;
      btn5ColorOn1 : String[10];   // enter: red OR green OR blue OR yellow OR white OR off
      btn5ColorOn2 : String[10];
      btn5ColorOff : String[10];   // enter: red OR green OR blue OR yellow OR white OR off
      btn6Activate : Bool;   // true for on, false for off
      btn6Mode : Bool;   // true for maintained, false for momentary
      btn6Group : Int;
      btn6Flash : Bool;
      btn6ColorOn1 : String[10];   // enter: red OR green OR blue OR yellow OR white OR off
      btn6ColorOn2 : String[10];
      btn6ColorOff : String[10];   // enter: red OR green OR blue OR yellow OR white OR off
      btn7Activate : Bool;   // true for on, false for off
      btn7Mode : Bool;   // true for maintained, false for momentary
      btn7Group : Int;
      btn7Flash : Bool;
      btn7ColorOn1 : String[10];   // enter: red OR green OR blue OR yellow OR white OR off
      btn7ColorOn2 : String[10];
      btn7ColorOff : String[10];   // enter: red OR green OR blue OR yellow OR white OR off
   END_VAR
   VAR_OUTPUT
      btnStatesOut : Array[0..7] of Bool;   // the output array represents the state of button presses
      btnColorsOut : DWord;
   END_VAR
   VAR
      mask : Byte;
      btnInInt : Byte;
      btnEval : Byte;
      i1 : Int;
      i2 : Int;
      btnActivateInt : Array[0..7] of Bool;
      btnClrMskOffInt : Array[0..7] of DWord;
      btnClrMskOn1Int : Array[0..7] of DWord;
      btnClrMskOn2Int : Array[0..7] of DWord;
      btnClrOffInt : Array[0..7] of String[10];
      btnClrOn1Int : Array[0..7] of String[10];
      btnClrOn2Int : Array[0..7] of String[10];
      btnColors : DWord;
      btnInArrayNew : Array[0..7] of Bool;
      btnInArrayOld : Array[0..7] of Bool;
      btnStateArrayInt : Array[0..7] of Bool;
      btnModeInt : Array[0..7] of Bool;
      btnFlashInt : Array[0..7] of Bool;
      btnGroup : Array[0..7] of Int;
   END_VAR
   VAR CONSTANT
      btnMskRed : DWord := dw#16#0100_0000;
      btnMskGreen : DWord := dw#16#0001_0000;
      btnMskBlue : DWord := dw#16#000_0100;
      btnMskYellow : DWord := dw#16#0101_0000;
      btnMskWhite : DWord := dw#16#0101_0100;
      btnMskBlack : DWord := dw#16#FEFE_FEFF;
      initBtnColors : DWord := dw#16#0000_0000;
   END_VAR
BEGIN
   REGION "ALL INITS"
       IF #hardInit OR #softInit THEN

           REGION "CLEAR OUTPUT COLORS"
               #btnColors := #initBtnColors;
           END_REGION

           REGION "TRANSFER PARAMETERS TO INTERNAL ARRAYS"

               REGION "BUTTON 0"
                   #btnActivateInt[0] := #btn0Activate;
                   #btnModeInt[0] := #btn0Mode;
                   #btnGroup[0] := #btn0Group;
                   #btnClrOn1Int[0] := #btn0ColorOn1;
                   #btnClrOn2Int[0] := #btn0ColorOn2;
                   #btnClrOffInt[0] := #btn0ColorOff;
               END_REGION

               REGION "BUTTON 1"
                   #btnActivateInt[1] := #btn1Activate;
                   #btnModeInt[1] := #btn1Mode;
                   #btnGroup[1] := #btn1Group;
                   #btnClrOn1Int[1] := #btn1ColorOn1;
                   #btnClrOn2Int[1] := #btn1ColorOn2;
                   #btnClrOffInt[1] := #btn1ColorOff;
               END_REGION

               REGION "BUTTON 2"
                   #btnActivateInt[2] := #btn2Activate;
                   #btnModeInt[2] := #btn2Mode;
                   #btnGroup[2] := #btn2Group;
                   #btnClrOn1Int[2] := #btn2ColorOn1;
                   #btnClrOn2Int[2] := #btn2ColorOn2;
                   #btnClrOffInt[2] := #btn2ColorOff;
               END_REGION

